// TIA Portal project "ROLLINGMILLPLC" (V16)

(* hardware
DEVICE "S71500/ET200MP station_1"  S7-1500 station
   slot 0: "Rail_0"  Rack  6ES7 590-1***0-0AA0
   slot 1: "PLC_1"  CPU 1518-4 PN/DP MFP  6ES7 518-4AX00-1AB0  V2.8
      slot 3: "CPU display_1"  6ES7591-1BA00-0AA0
      slot 32768: "PROFINET interface_1"  X1
         slot 32769: "Port_1"  X1 P1
         slot 32770: "Port_2"  X1 P2
      slot 33024: "PROFINET interface_2"  X2
         slot 33025: "Port_1"  X2 P1
      slot 33280: "PROFINET interface GBIT_3"  X3
         slot 33281: "Port_1"  X3 P1
      slot 33536: "DP interface_1"  X4
      slot 34817: "Virtual CP interface port_1"  Virtual CP interface port  Virtual CP interface port
DEVICE "S71500/ET200MP station_2"  S7-1500 station
   slot 0: "Rail_0"  Rack  6ES7 590-1***0-0AA0
   slot 1: "PLC_2"  CPU 1518-4 PN/DP MFP  6ES7 518-4AX00-1AB0  V2.8
      slot 3: "CPU display_1"  6ES7591-1BA00-0AA0
      slot 32768: "PROFINET interface_1"  X1
         slot 32769: "Port_1"  X1 P1
         slot 32770: "Port_2"  X1 P2
      slot 33024: "PROFINET interface_2"  X2
         slot 33025: "Port_1"  X2 P1
      slot 33280: "PROFINET interface GBIT_3"  X3
         slot 33281: "Port_1"  X3 P1
      slot 33536: "DP interface_1"  X4
      slot 34817: "Virtual CP interface port_1"  Virtual CP interface port  Virtual CP interface port
DEVICE "S71500/ET200MP station_3"  S7-1500 station
   slot 0: "Rail_0"  Rack  6ES7 590-1***0-0AA0
   slot 1: "PLC_3"  CPU 1518-4 PN/DP MFP  6ES7 518-4AX00-1AB0  V2.8
      slot 3: "CPU display_1"  6ES7591-1BA00-0AA0
      slot 32768: "PROFINET interface_1"  X1
         slot 32769: "Port_1"  X1 P1
         slot 32770: "Port_2"  X1 P2
      slot 33024: "PROFINET interface_2"  X2
         slot 33025: "Port_1"  X2 P1
      slot 33280: "PROFINET interface GBIT_3"  X3
         slot 33281: "Port_1"  X3 P1
      slot 33536: "DP interface_1"  X4
      slot 34817: "Virtual CP interface port_1"  Virtual CP interface port  Virtual CP interface port
DEVICE "HMI"  TP1500 Comfort
   slot 0: "HMI"  TP1500 Comfort  6AV2 124-0QC02-0AX0  16.0.0.0
   slot 1: "HMI_RT_2"  TP1500 Comfort  6AV2 124-0QC02-0AX0  16.0.0.0
   slot 5: "HMI.IE_CP_1"  PROFINET Interface  16.0.0.0
      slot 1: "PROFINET Interface_1"  PROFINET Interface
         slot 1: "Port_1"  Port
         slot 2: "Port_2"  Port
   slot 6: "HMI.IE_CP_2"  PROFINET Interface  16.0.0.0
      slot 1: "PROFINET Interface_GBit"  PROFINET Interface
         slot 1: "Port_1"  Port
   slot 7: "HMI.MPI/DP_CP_1"  MPI/DP Interface  16.0.0.0
*)

// ===== PLC "PLC_1"  CPU 1518-4 PN/DP MFP =====

TYPE "LQInternalModelSignals"
// This block is AUTO GENERATED - DO NOT MODIFY this block!
// Created by ODK_CodeGenerator version 205.100.101.18
// at Fri August 27 01:27:48 2021
// ********************************************************
   STRUCT
      Controlinput : Array[0..1] of LReal;
      Feedback : Array[0..4] of LReal;
      LQ_Refthickness : LReal;
      LQ_Refrollingforce : LReal;
   END_STRUCT;
END_TYPE

TYPE "LQParams"
// This block is AUTO GENERATED - DO NOT MODIFY this block!
// Created by ODK_CodeGenerator version 205.100.101.18
// at Mon August 30 17:02:50 2021
// ********************************************************
   STRUCT
      Lr : Array[0..3] of LReal;   // [LQ Controller 1/Gain Lr]:LQ_P.Lr
      Ly : Array[0..9] of LReal;   // [LQ Controller 1/Gain Ly]:LQ_P.Ly
   END_STRUCT;
   // Lr[0] := 0.013106;
   // Lr[1] := 0.0;
   // Lr[2] := 0.0;
   // Lr[3] := 3.112673;
   // Ly[0] := 0.0;
   // Ly[1] := 0.0;
   // Ly[2] := 0.0;
   // Ly[3] := 0.0;
   // Ly[4] := 0.011684;
   // Ly[5] := 0.0;
   // Ly[6] := 3.8E-05;
   // Ly[7] := 0.0;
   // Ly[8] := 0.0;
   // Ly[9] := 3.112673;
END_TYPE

DATA_BLOCK "LQ_GlobalData"   // DB1
{ S7_Optimized_Access := 'TRUE' }
VERSION : 0.1
   VAR
      Parameters : Struct
         thicknes : LReal;
         force : LReal;
      END_STRUCT;
      Feedback : Array[0..4] of LReal;
      Controlinput : Struct
         xv : LReal;
         fx : LReal;
      END_STRUCT;
      InternalModelSignals : "LQInternalModelSignals";
   END_VAR
   VAR RETAIN
      Param : "LQParams";
   END_VAR
BEGIN
END_DATA_BLOCK

DATA_BLOCK "gDB_SWV_Interface"   // DB2
{ S7_Optimized_Access := 'TRUE' }
VERSION : 0.1
// stored: InstanceOfName LQWebReadWrite
"LQWebReadWrite"
BEGIN
END_DATA_BLOCK

DATA_BLOCK "LQ_Unload_DB"   // DB3
{ S7_Optimized_Access := 'TRUE' }
VERSION : 0.1
// stored: InstanceOfName LQ_Unload
"LQ_Unload"
BEGIN
END_DATA_BLOCK

DATA_BLOCK "LQ_Load_DB"   // DB4
{ S7_Optimized_Access := 'TRUE' }
VERSION : 0.1
// stored: InstanceOfName LQ_Load
"LQ_Load"
BEGIN
END_DATA_BLOCK

DATA_BLOCK "LQOneStep_DB"   // DB5
{ S7_Optimized_Access := 'TRUE' }
VERSION : 0.1
// stored: InstanceOfName LQOneStep
"LQOneStep"
BEGIN
END_DATA_BLOCK

DATA_BLOCK "LQReadWriteParameters_DB"   // DB6
{ S7_Optimized_Access := 'TRUE' }
VERSION : 0.1
// stored: InstanceOfName LQReadWriteParameters
"LQReadWriteParameters"
BEGIN
END_DATA_BLOCK

DATA_BLOCK "OpcInterface"   // DB7
{ S7_Optimized_Access := 'TRUE' }
VERSION : 0.1
   VAR
      Feedback : Array[0..4] of LReal;
      Controlinput : Struct
         xv : LReal;
         fx : LReal;
      END_STRUCT;
   END_VAR
BEGIN
END_DATA_BLOCK

FUNCTION_BLOCK "LQ_Load"   // FB1, SCL
{ S7_Optimized_Access := 'TRUE' }
VERSION : 0.1
// This block is AUTO GENERATED - DO NOT MODIFY this block!
// Created by ODK_CodeGenerator version 2.5.1
// at Fri August 27 01:27:48 2021
// max. number of parallel calls into this ODK application is: 1
// *************************************************************
   VAR_INPUT
      REQ : Bool;
   END_VAR
   VAR_OUTPUT
      DONE : Bool;
      BUSY : Bool;
      ERROR : Bool;
      STATUS : Int;
   END_VAR
   VAR
      ODK_Load_Instance : ODK_Load;
      _odk_internal_LIBRARY_NAME : String := '<rt>LQ_ODK.so';
   END_VAR
   VAR CONSTANT
      _odk_internal_INSTANCE_ID : UDInt := 2_165_467_194;
   END_VAR
BEGIN
   //
   // DO NOT CHANGE BELOW OF THIS LINE !!
   // This is an automatic generated block by the
   // SIMATIC ODK 1500S V2.5.1
   // DO NOT CHANGE !!
   //
   #ODK_Load_Instance(REQ := #REQ,
                      LIBRARY_NAME := #_odk_internal_LIBRARY_NAME,
                      INSTANCE_ID := #_odk_internal_INSTANCE_ID,
                      DONE => #DONE,
                      BUSY => #BUSY,
                      ERROR => #ERROR,
                      STATUS => #STATUS);
   //
   // DO NOT CHANGE !!
   // This is an automatic generated block by the
   // SIMATIC ODK 1500S V2.5.1
   // DO NOT CHANGE ABOVE OF THIS LINE !!
   //
END_FUNCTION_BLOCK

FUNCTION_BLOCK "LQ_Unload"   // FB2, SCL
{ S7_Optimized_Access := 'TRUE' }
VERSION : 0.1
// This block is AUTO GENERATED - DO NOT MODIFY this block!
// Created by ODK_CodeGenerator version 205.100.101.18
// at Fri August 27 01:27:48 2021
// max. number of parallel calls into this ODK application is: 1
// *************************************************************
   VAR_INPUT
      REQ : Bool;
   END_VAR
   VAR_OUTPUT
      DONE : Bool;
      BUSY : Bool;
      ERROR : Bool;
      STATUS : Int;
   END_VAR
   VAR
      ODK_Unld_Instance : ODK_Unld;
   END_VAR
   VAR CONSTANT
      _odk_internal_INSTANCE_ID : UDInt := 2_165_467_194;
   END_VAR
BEGIN
   //
   // DO NOT CHANGE BELOW OF THIS LINE !!
   // This is an automatic generated block by the
   // SIMATIC ODK 1500S V2.5.1
   // DO NOT CHANGE !!
   //
   #ODK_Unld_Instance(REQ := #REQ,
                      INSTANCE_ID := #_odk_internal_INSTANCE_ID,
                      DONE => #DONE,
                      BUSY => #BUSY,
                      ERROR => #ERROR,
                      STATUS => #STATUS);
   //
   // DO NOT CHANGE !!
   // This is an automatic generated block by the
   // SIMATIC ODK 1500S V2.5.1
   // DO NOT CHANGE ABOVE OF THIS LINE !!
   //
END_FUNCTION_BLOCK

FUNCTION_BLOCK "LQOneStep"   // FB3, SCL
{ S7_Optimized_Access := 'TRUE' }
VERSION : 0.1
// This block is AUTO GENERATED - DO NOT MODIFY this block!
// Created by ODK_CodeGenerator version 205.100.101.18
// at Fri August 27 01:27:48 2021
// max. number of parallel calls into this ODK application is: 1
// *************************************************************
//  This is generated by Target 1500S for Simulink
//  Model name:                  LQ
//  Model version:               1.16
//                 
//  ODK 1500S version:           V2.5
//  Target 1500S version:        V4.0         
//  MATLAB version:              9.9 (R2020b) 29-Jul-2020
//  Simulink version:            10.2 (R2020b) 29-Jul-2020
//  MATLAB Coder version:        5.1 (R2020b) 29-Jul-2020
//  Simulink Coder version:      9.4 (R2020b) 29-Jul-2020
//  
//  ***Model details***
//  Step Size:                   0.01
//  Default parameter behaviour: Tunable
//  External Mode:               Off
//  
//  ***ODK 1500S details***  
//  Heap Size:                   32k
//  Max Block Size:              1024
//  Size of thread stack:        32k
//  SyncCallParallelCount:       1(max. number of parallel calls into this ODK application)
//  ********************************************************
   VAR_INPUT
      Feedback : Array[0..4] of LReal;
      Refthickness : LReal;
      Refrollingforce : LReal;
   END_VAR
   VAR_OUTPUT
      STATUS : Int := 0;
      xv : LReal;
      fx : LReal;
      internalSignals : "LQInternalModelSignals";
   END_VAR
   VAR
      _odk_internal_Last_REQ : Bool := FALSE;
      _odk_internal_Last_BUSY : Bool := FALSE;
      _odk_internal_IN_BUFFER : Array[0..55] of Byte;
      _odk_internal_OUT_BUFFER : Array[0..87] of Byte;
   END_VAR
   VAR_TEMP
      _odk_internal_pos : DInt;
      _odk_internal_err : Int;
      _odk_internal_i : Int;
   END_VAR
   VAR CONSTANT
      _odk_internal_INSTANCE_ID : UDInt := 2_165_467_194;
      _odk_internal_COMMAND : UDInt := 295_977_560;
   END_VAR
BEGIN
   //
   // DO NOT CHANGE BELOW OF THIS LINE !!
   // This is an automatic generated block by the
   // SIMATIC ODK 1500S V2.5.1
   // DO NOT CHANGE !!
   //
   // This is generated by Target 1500S for Simulink
   // Model name:                  LQ
   // Model version:               1.16
   //                
   // ODK 1500S version:           V2.5
   // Target 1500S version:        V4.0         
   // MATLAB version:              9.9 (R2020b) 29-Jul-2020
   // Simulink version:            10.2 (R2020b) 29-Jul-2020
   // MATLAB Coder version:        5.1 (R2020b) 29-Jul-2020
   // Simulink Coder version:      9.4 (R2020b) 29-Jul-2020
   // 
   // ***Model details***
   // Step Size:                   0.01
   // Default parameter behaviour: Tunable
   // External Mode:               Off
   // 
   // ***ODK 1500S details***  
   // Heap Size:                   32k
   // Max Block Size:              1024
   // Size of thread stack:        32k
   // SyncCallParallelCount:       1(max. number of parallel calls into this ODK application)
   // ********************************************************
   // 
   #_odk_internal_pos := 0;
   FOR #_odk_internal_i := 0 TO 4 DO
       #_odk_internal_err := WRITE_LITTLE(src_variable := #Feedback[#_odk_internal_i], dest_array := #_odk_internal_IN_BUFFER, pos := #_odk_internal_pos);
   END_FOR;
   #_odk_internal_err := WRITE_LITTLE(src_variable := #Refthickness, dest_array := #_odk_internal_IN_BUFFER, pos := #_odk_internal_pos);
   #_odk_internal_err := WRITE_LITTLE(src_variable := #Refrollingforce, dest_array := #_odk_internal_IN_BUFFER, pos := #_odk_internal_pos);
   #STATUS := ODK_ExcS(INSTANCE_ID := #_odk_internal_INSTANCE_ID,
                       COMMAND := #_odk_internal_COMMAND,
                       IN_DATA := #_odk_internal_IN_BUFFER,
                       INOUT_DATA := null,
                       OUT_DATA := #_odk_internal_OUT_BUFFER
   );
   IF INT_TO_UINT(#STATUS) < 16#7000 THEN
       #_odk_internal_pos := 0;
       #_odk_internal_err := READ_LITTLE(dest_Variable => #xv, src_array := #_odk_internal_OUT_BUFFER, pos := #_odk_internal_pos);
       #_odk_internal_err := READ_LITTLE(dest_Variable => #fx, src_array := #_odk_internal_OUT_BUFFER, pos := #_odk_internal_pos);
       FOR #_odk_internal_i := 0 TO 1 DO
           #_odk_internal_err := READ_LITTLE(dest_Variable => #internalSignals.#Controlinput[#_odk_internal_i], src_array := #_odk_internal_OUT_BUFFER, pos := #_odk_internal_pos);
       END_FOR;
       FOR #_odk_internal_i := 0 TO 4 DO
           #_odk_internal_err := READ_LITTLE(dest_Variable => #internalSignals.#Feedback[#_odk_internal_i], src_array := #_odk_internal_OUT_BUFFER, pos := #_odk_internal_pos);
       END_FOR;
       #_odk_internal_err := READ_LITTLE(dest_Variable => #internalSignals.#LQ_Refthickness, src_array := #_odk_internal_OUT_BUFFER, pos := #_odk_internal_pos);
       #_odk_internal_err := READ_LITTLE(dest_Variable => #internalSignals.#LQ_Refrollingforce, src_array := #_odk_internal_OUT_BUFFER, pos := #_odk_internal_pos);
   END_IF;
   //
   // DO NOT CHANGE !!
   // This is an automatic generated block by the
   // SIMATIC ODK 1500S V2.5.1
   // DO NOT CHANGE ABOVE OF THIS LINE !!
   //
END_FUNCTION_BLOCK

FUNCTION_BLOCK "LQReadWriteParameters"   // FB4, SCL
{ S7_Optimized_Access := 'TRUE' }
VERSION : 0.1
// This block is AUTO GENERATED - DO NOT MODIFY this block!
// Created by ODK_CodeGenerator version 205.100.101.18
// at Fri August 27 01:27:49 2021
// max. number of parallel calls into this ODK application is: 1
// *************************************************************
//  This is generated by Target 1500S for Simulink
//  Model name:                  LQ
//  Model version:               1.16
//                 
//  ODK 1500S version:           V2.5
//  Target 1500S version:        V4.0         
//  MATLAB version:              9.9 (R2020b) 29-Jul-2020
//  Simulink version:            10.2 (R2020b) 29-Jul-2020
//  MATLAB Coder version:        5.1 (R2020b) 29-Jul-2020
//  Simulink Coder version:      9.4 (R2020b) 29-Jul-2020
//  
//  ***Model details***
//  Step Size:                   0.01
//  Default parameter behaviour: Tunable
//  External Mode:               Off
//  
//  ***ODK 1500S details***  
//  Heap Size:                   32k
//  Max Block Size:              1024
//  Size of thread stack:        32k
//  SyncCallParallelCount:       1(max. number of parallel calls into this ODK application)
//  ********************************************************
//  
//  Call this function to read or write parameters from/to Simulink Model.
//  Set write[IN] parameter to TRUE in order to write and set FALSE to read parameters
   VAR_INPUT
      write : Bool;
   END_VAR
   VAR_OUTPUT
      STATUS : Int := 0;
   END_VAR
   VAR_IN_OUT
      inOutParams : "LQParams";
   END_VAR
   VAR
      _odk_internal_Last_REQ : Bool := FALSE;
      _odk_internal_Last_BUSY : Bool := FALSE;
      _odk_internal_IN_BUFFER : Array[0..0] of Byte;
      _odk_internal_INOUT_BUFFER : Array[0..111] of Byte;
   END_VAR
   VAR_TEMP
      _odk_internal_pos : DInt;
      _odk_internal_err : Int;
      _odk_internal_i : Int;
   END_VAR
   VAR CONSTANT
      _odk_internal_INSTANCE_ID : UDInt := 2_165_467_194;
      _odk_internal_COMMAND : UDInt := 2_137_970_399;
   END_VAR
BEGIN
   //
   // DO NOT CHANGE BELOW OF THIS LINE !!
   // This is an automatic generated block by the
   // SIMATIC ODK 1500S V2.5.1
   // DO NOT CHANGE !!
   //
   // This is generated by Target 1500S for Simulink
   // Model name:                  LQ
   // Model version:               1.16
   //                
   // ODK 1500S version:           V2.5
   // Target 1500S version:        V4.0         
   // MATLAB version:              9.9 (R2020b) 29-Jul-2020
   // Simulink version:            10.2 (R2020b) 29-Jul-2020
   // MATLAB Coder version:        5.1 (R2020b) 29-Jul-2020
   // Simulink Coder version:      9.4 (R2020b) 29-Jul-2020
   // 
   // ***Model details***
   // Step Size:                   0.01
   // Default parameter behaviour: Tunable
   // External Mode:               Off
   // 
   // ***ODK 1500S details***  
   // Heap Size:                   32k
   // Max Block Size:              1024
   // Size of thread stack:        32k
   // SyncCallParallelCount:       1(max. number of parallel calls into this ODK application)
   // ********************************************************
   // 
   // Call this function to read or write parameters from/to Simulink Model.
   // Set write[IN] parameter to TRUE in order to write and set FALSE to read parameters
   #_odk_internal_pos := 0;
   IF (True = #write) THEN
       #_odk_internal_IN_BUFFER[#_odk_internal_pos] := BYTE#1;
   ELSE
       #_odk_internal_IN_BUFFER[#_odk_internal_pos] := BYTE#0;
   END_IF;
   #_odk_internal_pos := #_odk_internal_pos + 1;
   #_odk_internal_pos := 0;
   FOR #_odk_internal_i := 0 TO 3 DO
       #_odk_internal_err := WRITE_LITTLE(src_variable := #inOutParams.#Lr[#_odk_internal_i], dest_array := #_odk_internal_INOUT_BUFFER, pos := #_odk_internal_pos);
   END_FOR;
   FOR #_odk_internal_i := 0 TO 9 DO
       #_odk_internal_err := WRITE_LITTLE(src_variable := #inOutParams.#Ly[#_odk_internal_i], dest_array := #_odk_internal_INOUT_BUFFER, pos := #_odk_internal_pos);
   END_FOR;
   #STATUS := ODK_ExcS(INSTANCE_ID := #_odk_internal_INSTANCE_ID,
                       COMMAND := #_odk_internal_COMMAND,
                       IN_DATA := #_odk_internal_IN_BUFFER,
                       INOUT_DATA := #_odk_internal_INOUT_BUFFER,
                       OUT_DATA := null);
   IF INT_TO_UINT(#STATUS) < 16#7000 THEN
       #_odk_internal_pos := 0;
       FOR #_odk_internal_i := 0 TO 3 DO
           #_odk_internal_err := READ_LITTLE(dest_Variable => #inOutParams.#Lr[#_odk_internal_i], src_array := #_odk_internal_INOUT_BUFFER, pos := #_odk_internal_pos);
       END_FOR;
       FOR #_odk_internal_i := 0 TO 9 DO
           #_odk_internal_err := READ_LITTLE(dest_Variable => #inOutParams.#Ly[#_odk_internal_i], src_array := #_odk_internal_INOUT_BUFFER, pos := #_odk_internal_pos);
       END_FOR;
   END_IF;
   //
   // DO NOT CHANGE !!
   // This is an automatic generated block by the
   // SIMATIC ODK 1500S V2.5.1
   // DO NOT CHANGE ABOVE OF THIS LINE !!
   //
END_FUNCTION_BLOCK

FUNCTION_BLOCK "LQWebReadWrite"   // FB5, SCL
{ S7_Optimized_Access := 'TRUE' }
VERSION : 0.1
// This block is AUTO GENERATED - DO NOT MODIFY this block!
// Created by Target 1500S version 0
// at 0 
// ********************************************************
//  This is generated by Target 1500S for Simulink
//  Model name:                  LQ
//  Model version:               1.16
//                
//  ODK 1500S version:           V2.5
//  Target 1500S version:        V4.0         
//  MATLAB version:              9.9 (R2020b) 29-Jul-2020
//  Simulink version:            10.2 (R2020b) 29-Jul-2020
//  MATLAB Coder version:        5.1 (R2020b) 29-Jul-2020
//  Simulink Coder version:      9.4 (R2020b) 29-Jul-2020
// 
//  ***Model details***
//  Step Size:                   0.01
//  Default parameter behaviour: Tunable 
//  External Mode:               Off
//  ***ODK 1500S details***  
//  Heap Size:                   32k
//  Max Block Size:              1024
//  Size of thread stack:        32k
//  SyncCallParallelCount:       1(max. number of parallel calls into this ODK application)
//  ********************************************************
// Call this FB to establish a connection to user defined Web page.
   VAR_INPUT
      InternalSignals : "LQInternalModelSignals";
      CTRL_DB : DB_WWW;
   END_VAR
   VAR_IN_OUT
      Params : "LQParams";
   END_VAR
   VAR
      TestPointedSignals : "LQInternalModelSignals";
      Parameter : "LQParams";
      RWParams_Instance : "LQReadWriteParameters";
      Write : Int := 0;
      RunTime : LReal;
   END_VAR
   VAR_TEMP
      ret : Int;
   END_VAR
BEGIN
   // This is generated by Target 1500S for Simulink
   // Model name:                  LQ
   // Model version:               1.16
   //               
   // ODK 1500S version:           V2.5
   // Target 1500S version:        V4.0         
   // MATLAB version:              9.9 (R2020b) 29-Jul-2020
   // Simulink version:            10.2 (R2020b) 29-Jul-2020
   // MATLAB Coder version:        5.1 (R2020b) 29-Jul-2020
   // Simulink Coder version:      9.4 (R2020b) 29-Jul-2020
   //
   // ***Model details***
   // Step Size:                   0.01
   // Default parameter behaviour: Tunable 
   // External Mode:               Off
   // ***ODK 1500S details***  
   // Heap Size:                   32k
   // Max Block Size:              1024
   // Size of thread stack:        32k
   // SyncCallParallelCount:       1(max. number of parallel calls into this ODK application)
   // ********************************************************
   //Call this FB to establish a connection to user defined Web page.
   #RunTime := #RunTime + 10.0;

   #TestPointedSignals := #InternalSignals;
   CASE #Write OF
       0:
           #RWParams_Instance(write := FALSE,
                              STATUS => #RWParams_Instance.STATUS,
                              inOutParams := #Parameter);
           #Params := #Parameter;
       1:
           // Wait for parameter be updated by the Web action
           ;
       2:
           #RWParams_Instance(write := TRUE,
                              STATUS => #RWParams_Instance.STATUS,
                              inOutParams := #Parameter);
           #Params := #Parameter;
           #Write := 0;
       ELSE
           // Not possible to reach
           ;
   END_CASE;

   #ret := WWW(#CTRL_DB);
END_FUNCTION_BLOCK

ORGANIZATION_BLOCK "Main"   // OB1, LAD, ProgramCycle
TITLE = "Main Program Sweep (Cycle)"
{ S7_Optimized_Access := 'TRUE' }
VERSION : 0.1
   VAR_INPUT
      Initial_Call : Bool;   // Initial call of this OB
      Remanence : Bool;   // =True, if remanent data are available
   END_VAR
BEGIN
END_ORGANIZATION_BLOCK

ORGANIZATION_BLOCK "Cyclic interrupt"   // OB30, LAD, CyclicInterrupt
{ S7_Optimized_Access := 'TRUE' }
VERSION : 0.1
   VAR_INPUT
      Initial_Call : Bool;   // Initial call of this OB
      Event_Count : Int;   // Events discarded
   END_VAR
BEGIN

REGION Network 1 (SCL)
   "LQ_GlobalData".Feedback := "OpcInterface".Feedback;
END_REGION

REGION Network 2
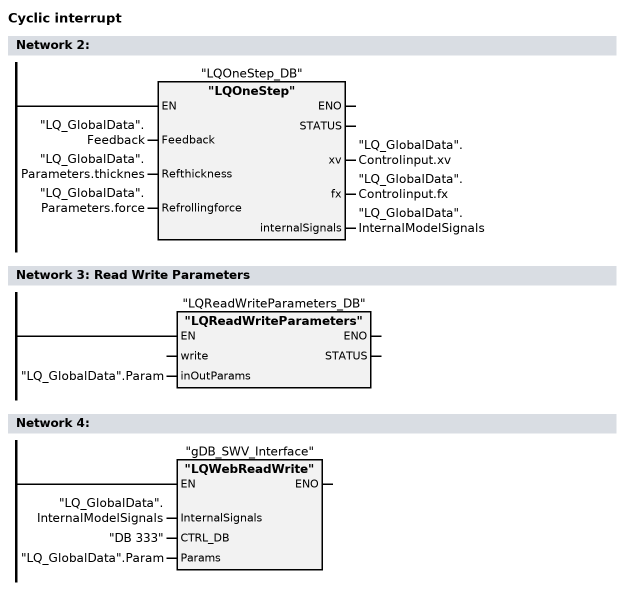
   RUNG wire#powerrail
      "LQOneStep_DB"(Feedback := "LQ_GlobalData".Feedback, Refthickness := "LQ_GlobalData".Parameters.thicknes, Refrollingforce := "LQ_GlobalData".Parameters.force, STATUS =>, xv => "LQ_GlobalData".Controlinput.xv, fx => "LQ_GlobalData".Controlinput.fx, internalSignals => "LQ_GlobalData".InternalModelSignals)
   END_RUNG
   // the same network as SCL:
   "LQOneStep_DB"(Feedback := "LQ_GlobalData".Feedback,   // "LQOneStep"
                  Refthickness := "LQ_GlobalData".Parameters.thicknes,
                  Refrollingforce := "LQ_GlobalData".Parameters.force,
                  xv => "LQ_GlobalData".Controlinput.xv,
                  fx => "LQ_GlobalData".Controlinput.fx,
                  internalSignals => "LQ_GlobalData".InternalModelSignals);
END_REGION

REGION Network 3: Read Write Parameters
   RUNG wire#powerrail
      "LQReadWriteParameters_DB"(write :=, inOutParams := "LQ_GlobalData".Param, STATUS =>)
   END_RUNG
   // the same network as SCL:
   "LQReadWriteParameters_DB"(inOutParams := "LQ_GlobalData".Param);   // "LQReadWriteParameters"
END_REGION

REGION Network 4
   RUNG wire#powerrail
      "gDB_SWV_Interface"(InternalSignals := "LQ_GlobalData".InternalModelSignals, CTRL_DB := "DB 333", Params := "LQ_GlobalData".Param)
   END_RUNG
   // the same network as SCL:
   "gDB_SWV_Interface"(InternalSignals := "LQ_GlobalData".InternalModelSignals,   // "LQWebReadWrite"
                       CTRL_DB := "DB 333",
                       Params := "LQ_GlobalData".Param);
END_REGION

REGION Network 5 (SCL)
   "OpcInterface".Controlinput.xv := "LQ_GlobalData".Controlinput.xv;
   "OpcInterface".Controlinput.fx := "LQ_GlobalData".Controlinput.fx;
END_REGION
END_ORGANIZATION_BLOCK

ORGANIZATION_BLOCK "Startup"   // OB100, LAD, Startup
TITLE = "Complete Restart"
{ S7_Optimized_Access := 'TRUE' }
VERSION : 0.1
   VAR_INPUT
      LostRetentive : Bool;   // True if retentive data are lost
      LostRTC : Bool;   // True if date and time are lost
   END_VAR
BEGIN

REGION Network 1
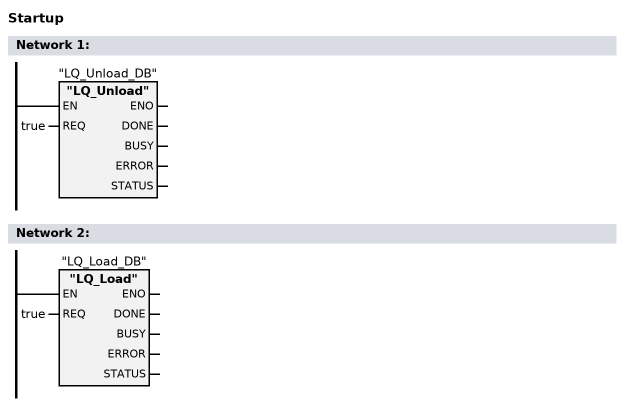
   RUNG wire#powerrail
      "LQ_Unload_DB"(REQ := true, DONE =>, BUSY =>, ERROR =>, STATUS =>)
   END_RUNG
   // the same network as SCL:
   "LQ_Unload_DB"(REQ := true);   // "LQ_Unload"
END_REGION

REGION Network 2
   RUNG wire#powerrail
      "LQ_Load_DB"(REQ := true, DONE =>, BUSY =>, ERROR =>, STATUS =>)
   END_RUNG
   // the same network as SCL:
   "LQ_Load_DB"(REQ := true);   // "LQ_Load"
END_REGION
END_ORGANIZATION_BLOCK

// ===== PLC "PLC_2"  CPU 1518-4 PN/DP MFP =====

TYPE "LQInternalModelSignals"
// This block is AUTO GENERATED - DO NOT MODIFY this block!
// Created by ODK_CodeGenerator version 205.100.101.18
// at Fri August 27 01:31:13 2021
// ********************************************************
   STRUCT
      Controlinput : Array[0..1] of LReal;
      Feedback : Array[0..4] of LReal;
      LQ_Refthickness : LReal;
      LQ_Refrollingforce : LReal;
   END_STRUCT;
END_TYPE

TYPE "LQParams"
// This block is AUTO GENERATED - DO NOT MODIFY this block!
// Created by ODK_CodeGenerator version 205.100.101.18
// at Mon August 30 17:02:50 2021
// ********************************************************
   STRUCT
      Lr : Array[0..3] of LReal;   // [LQ Controller 1/Gain Lr]:LQ_P.Lr
      Ly : Array[0..9] of LReal;   // [LQ Controller 1/Gain Ly]:LQ_P.Ly
   END_STRUCT;
   // Lr[0] := 0.013106;
   // Lr[1] := 0.0;
   // Lr[2] := 0.0;
   // Lr[3] := 3.112673;
   // Ly[0] := 0.0;
   // Ly[1] := 0.0;
   // Ly[2] := 0.0;
   // Ly[3] := 0.0;
   // Ly[4] := 0.011684;
   // Ly[5] := 0.0;
   // Ly[6] := 3.8E-05;
   // Ly[7] := 0.0;
   // Ly[8] := 0.0;
   // Ly[9] := 3.112673;
END_TYPE

DATA_BLOCK "LQ_GlobalData"   // DB1
{ S7_Optimized_Access := 'TRUE' }
VERSION : 0.1
   VAR
      Parameters : Struct
         thicknes : LReal;
         force : LReal;
      END_STRUCT;
      Feedback : Array[0..4] of LReal;
      Controlinput : Struct
         xv : LReal;
         fx : LReal;
      END_STRUCT;
      InternalModelSignals : "LQInternalModelSignals";
   END_VAR
   VAR RETAIN
      Param : "LQParams";
   END_VAR
BEGIN
END_DATA_BLOCK

DATA_BLOCK "gDB_SWV_Interface"   // DB2
{ S7_Optimized_Access := 'TRUE' }
VERSION : 0.1
// stored: InstanceOfName LQWebReadWrite
"LQWebReadWrite"
BEGIN
END_DATA_BLOCK

DATA_BLOCK "OpcInterface"   // DB3
{ S7_Optimized_Access := 'TRUE' }
VERSION : 0.1
   VAR
      Feedback : Array[0..4] of LReal;
      Controlinput : Struct
         xv : LReal;
         fx : LReal;
      END_STRUCT;
   END_VAR
BEGIN
END_DATA_BLOCK

DATA_BLOCK "LQReadWriteParameters_DB"   // DB4
{ S7_Optimized_Access := 'TRUE' }
VERSION : 0.1
// stored: InstanceOfName LQReadWriteParameters
"LQReadWriteParameters"
BEGIN
END_DATA_BLOCK

DATA_BLOCK "LQ_Unload_DB"   // DB5
{ S7_Optimized_Access := 'TRUE' }
VERSION : 0.1
// stored: InstanceOfName LQ_Unload
"LQ_Unload"
BEGIN
END_DATA_BLOCK

DATA_BLOCK "LQOneStep_DB"   // DB7
{ S7_Optimized_Access := 'TRUE' }
VERSION : 0.1
// stored: InstanceOfName LQOneStep
"LQOneStep"
BEGIN
END_DATA_BLOCK

DATA_BLOCK "LQ_Load_DB"   // DB8
{ S7_Optimized_Access := 'TRUE' }
VERSION : 0.1
// stored: InstanceOfName LQ_Load
"LQ_Load"
BEGIN
END_DATA_BLOCK

FUNCTION_BLOCK "LQ_Load"   // FB1, SCL
{ S7_Optimized_Access := 'TRUE' }
VERSION : 0.1
// This block is AUTO GENERATED - DO NOT MODIFY this block!
// Created by ODK_CodeGenerator version 2.5.1
// at Fri August 27 01:31:13 2021
// max. number of parallel calls into this ODK application is: 1
// *************************************************************
   VAR_INPUT
      REQ : Bool;
   END_VAR
   VAR_OUTPUT
      DONE : Bool;
      BUSY : Bool;
      ERROR : Bool;
      STATUS : Int;
   END_VAR
   VAR
      ODK_Load_Instance : ODK_Load;
      _odk_internal_LIBRARY_NAME : String := '<rt>LQ_ODK.so';
   END_VAR
   VAR CONSTANT
      _odk_internal_INSTANCE_ID : UDInt := 2_363_350_554;
   END_VAR
BEGIN
   //
   // DO NOT CHANGE BELOW OF THIS LINE !!
   // This is an automatic generated block by the
   // SIMATIC ODK 1500S V2.5.1
   // DO NOT CHANGE !!
   //
   #ODK_Load_Instance(REQ := #REQ,
                      LIBRARY_NAME := #_odk_internal_LIBRARY_NAME,
                      INSTANCE_ID := #_odk_internal_INSTANCE_ID,
                      DONE => #DONE,
                      BUSY => #BUSY,
                      ERROR => #ERROR,
                      STATUS => #STATUS);
   //
   // DO NOT CHANGE !!
   // This is an automatic generated block by the
   // SIMATIC ODK 1500S V2.5.1
   // DO NOT CHANGE ABOVE OF THIS LINE !!
   //
END_FUNCTION_BLOCK

FUNCTION_BLOCK "LQ_Unload"   // FB2, SCL
{ S7_Optimized_Access := 'TRUE' }
VERSION : 0.1
// This block is AUTO GENERATED - DO NOT MODIFY this block!
// Created by ODK_CodeGenerator version 205.100.101.18
// at Fri August 27 01:31:13 2021
// max. number of parallel calls into this ODK application is: 1
// *************************************************************
   VAR_INPUT
      REQ : Bool;
   END_VAR
   VAR_OUTPUT
      DONE : Bool;
      BUSY : Bool;
      ERROR : Bool;
      STATUS : Int;
   END_VAR
   VAR
      ODK_Unld_Instance : ODK_Unld;
   END_VAR
   VAR CONSTANT
      _odk_internal_INSTANCE_ID : UDInt := 2_363_350_554;
   END_VAR
BEGIN
   //
   // DO NOT CHANGE BELOW OF THIS LINE !!
   // This is an automatic generated block by the
   // SIMATIC ODK 1500S V2.5.1
   // DO NOT CHANGE !!
   //
   #ODK_Unld_Instance(REQ := #REQ,
                      INSTANCE_ID := #_odk_internal_INSTANCE_ID,
                      DONE => #DONE,
                      BUSY => #BUSY,
                      ERROR => #ERROR,
                      STATUS => #STATUS);
   //
   // DO NOT CHANGE !!
   // This is an automatic generated block by the
   // SIMATIC ODK 1500S V2.5.1
   // DO NOT CHANGE ABOVE OF THIS LINE !!
   //
END_FUNCTION_BLOCK

FUNCTION_BLOCK "LQOneStep"   // FB3, SCL
{ S7_Optimized_Access := 'TRUE' }
VERSION : 0.1
// This block is AUTO GENERATED - DO NOT MODIFY this block!
// Created by ODK_CodeGenerator version 205.100.101.18
// at Fri August 27 01:31:13 2021
// max. number of parallel calls into this ODK application is: 1
// *************************************************************
//  This is generated by Target 1500S for Simulink
//  Model name:                  LQ
//  Model version:               1.16
//                 
//  ODK 1500S version:           V2.5
//  Target 1500S version:        V4.0         
//  MATLAB version:              9.9 (R2020b) 29-Jul-2020
//  Simulink version:            10.2 (R2020b) 29-Jul-2020
//  MATLAB Coder version:        5.1 (R2020b) 29-Jul-2020
//  Simulink Coder version:      9.4 (R2020b) 29-Jul-2020
//  
//  ***Model details***
//  Step Size:                   0.01
//  Default parameter behaviour: Tunable
//  External Mode:               Off
//  
//  ***ODK 1500S details***  
//  Heap Size:                   32k
//  Max Block Size:              1024
//  Size of thread stack:        32k
//  SyncCallParallelCount:       1(max. number of parallel calls into this ODK application)
//  ********************************************************
   VAR_INPUT
      Feedback : Array[0..4] of LReal;
      Refthickness : LReal;
      Refrollingforce : LReal;
   END_VAR
   VAR_OUTPUT
      STATUS : Int := 0;
      xv : LReal;
      fx : LReal;
      internalSignals : "LQInternalModelSignals";
   END_VAR
   VAR
      _odk_internal_Last_REQ : Bool := FALSE;
      _odk_internal_Last_BUSY : Bool := FALSE;
      _odk_internal_IN_BUFFER : Array[0..55] of Byte;
      _odk_internal_OUT_BUFFER : Array[0..87] of Byte;
   END_VAR
   VAR_TEMP
      _odk_internal_pos : DInt;
      _odk_internal_err : Int;
      _odk_internal_i : Int;
   END_VAR
   VAR CONSTANT
      _odk_internal_INSTANCE_ID : UDInt := 2_363_350_554;
      _odk_internal_COMMAND : UDInt := 295_977_560;
   END_VAR
BEGIN
   //
   // DO NOT CHANGE BELOW OF THIS LINE !!
   // This is an automatic generated block by the
   // SIMATIC ODK 1500S V2.5.1
   // DO NOT CHANGE !!
   //
   // This is generated by Target 1500S for Simulink
   // Model name:                  LQ
   // Model version:               1.16
   //                
   // ODK 1500S version:           V2.5
   // Target 1500S version:        V4.0         
   // MATLAB version:              9.9 (R2020b) 29-Jul-2020
   // Simulink version:            10.2 (R2020b) 29-Jul-2020
   // MATLAB Coder version:        5.1 (R2020b) 29-Jul-2020
   // Simulink Coder version:      9.4 (R2020b) 29-Jul-2020
   // 
   // ***Model details***
   // Step Size:                   0.01
   // Default parameter behaviour: Tunable
   // External Mode:               Off
   // 
   // ***ODK 1500S details***  
   // Heap Size:                   32k
   // Max Block Size:              1024
   // Size of thread stack:        32k
   // SyncCallParallelCount:       1(max. number of parallel calls into this ODK application)
   // ********************************************************
   // 
   #_odk_internal_pos := 0;
   FOR #_odk_internal_i := 0 TO 4 DO
       #_odk_internal_err := WRITE_LITTLE(src_variable := #Feedback[#_odk_internal_i], dest_array := #_odk_internal_IN_BUFFER, pos := #_odk_internal_pos);
   END_FOR;
   #_odk_internal_err := WRITE_LITTLE(src_variable := #Refthickness, dest_array := #_odk_internal_IN_BUFFER, pos := #_odk_internal_pos);
   #_odk_internal_err := WRITE_LITTLE(src_variable := #Refrollingforce, dest_array := #_odk_internal_IN_BUFFER, pos := #_odk_internal_pos);
   #STATUS := ODK_ExcS(INSTANCE_ID := #_odk_internal_INSTANCE_ID,
                       COMMAND := #_odk_internal_COMMAND,
                       IN_DATA := #_odk_internal_IN_BUFFER,
                       INOUT_DATA := null,
                       OUT_DATA := #_odk_internal_OUT_BUFFER
   );
   IF INT_TO_UINT(#STATUS) < 16#7000 THEN
       #_odk_internal_pos := 0;
       #_odk_internal_err := READ_LITTLE(dest_Variable => #xv, src_array := #_odk_internal_OUT_BUFFER, pos := #_odk_internal_pos);
       #_odk_internal_err := READ_LITTLE(dest_Variable => #fx, src_array := #_odk_internal_OUT_BUFFER, pos := #_odk_internal_pos);
       FOR #_odk_internal_i := 0 TO 1 DO
           #_odk_internal_err := READ_LITTLE(dest_Variable => #internalSignals.#Controlinput[#_odk_internal_i], src_array := #_odk_internal_OUT_BUFFER, pos := #_odk_internal_pos);
       END_FOR;
       FOR #_odk_internal_i := 0 TO 4 DO
           #_odk_internal_err := READ_LITTLE(dest_Variable => #internalSignals.#Feedback[#_odk_internal_i], src_array := #_odk_internal_OUT_BUFFER, pos := #_odk_internal_pos);
       END_FOR;
       #_odk_internal_err := READ_LITTLE(dest_Variable => #internalSignals.#LQ_Refthickness, src_array := #_odk_internal_OUT_BUFFER, pos := #_odk_internal_pos);
       #_odk_internal_err := READ_LITTLE(dest_Variable => #internalSignals.#LQ_Refrollingforce, src_array := #_odk_internal_OUT_BUFFER, pos := #_odk_internal_pos);
   END_IF;
   //
   // DO NOT CHANGE !!
   // This is an automatic generated block by the
   // SIMATIC ODK 1500S V2.5.1
   // DO NOT CHANGE ABOVE OF THIS LINE !!
   //
END_FUNCTION_BLOCK

FUNCTION_BLOCK "LQReadWriteParameters"   // FB4, SCL
{ S7_Optimized_Access := 'TRUE' }
VERSION : 0.1
// This block is AUTO GENERATED - DO NOT MODIFY this block!
// Created by ODK_CodeGenerator version 205.100.101.18
// at Fri August 27 01:31:13 2021
// max. number of parallel calls into this ODK application is: 1
// *************************************************************
//  This is generated by Target 1500S for Simulink
//  Model name:                  LQ
//  Model version:               1.16
//                 
//  ODK 1500S version:           V2.5
//  Target 1500S version:        V4.0         
//  MATLAB version:              9.9 (R2020b) 29-Jul-2020
//  Simulink version:            10.2 (R2020b) 29-Jul-2020
//  MATLAB Coder version:        5.1 (R2020b) 29-Jul-2020
//  Simulink Coder version:      9.4 (R2020b) 29-Jul-2020
//  
//  ***Model details***
//  Step Size:                   0.01
//  Default parameter behaviour: Tunable
//  External Mode:               Off
//  
//  ***ODK 1500S details***  
//  Heap Size:                   32k
//  Max Block Size:              1024
//  Size of thread stack:        32k
//  SyncCallParallelCount:       1(max. number of parallel calls into this ODK application)
//  ********************************************************
//  
//  Call this function to read or write parameters from/to Simulink Model.
//  Set write[IN] parameter to TRUE in order to write and set FALSE to read parameters
   VAR_INPUT
      write : Bool;
   END_VAR
   VAR_OUTPUT
      STATUS : Int := 0;
   END_VAR
   VAR_IN_OUT
      inOutParams : "LQParams";
   END_VAR
   VAR
      _odk_internal_Last_REQ : Bool := FALSE;
      _odk_internal_Last_BUSY : Bool := FALSE;
      _odk_internal_IN_BUFFER : Array[0..0] of Byte;
      _odk_internal_INOUT_BUFFER : Array[0..111] of Byte;
   END_VAR
   VAR_TEMP
      _odk_internal_pos : DInt;
      _odk_internal_err : Int;
      _odk_internal_i : Int;
   END_VAR
   VAR CONSTANT
      _odk_internal_INSTANCE_ID : UDInt := 2_363_350_554;
      _odk_internal_COMMAND : UDInt := 2_137_970_399;
   END_VAR
BEGIN
   //
   // DO NOT CHANGE BELOW OF THIS LINE !!
   // This is an automatic generated block by the
   // SIMATIC ODK 1500S V2.5.1
   // DO NOT CHANGE !!
   //
   // This is generated by Target 1500S for Simulink
   // Model name:                  LQ
   // Model version:               1.16
   //                
   // ODK 1500S version:           V2.5
   // Target 1500S version:        V4.0         
   // MATLAB version:              9.9 (R2020b) 29-Jul-2020
   // Simulink version:            10.2 (R2020b) 29-Jul-2020
   // MATLAB Coder version:        5.1 (R2020b) 29-Jul-2020
   // Simulink Coder version:      9.4 (R2020b) 29-Jul-2020
   // 
   // ***Model details***
   // Step Size:                   0.01
   // Default parameter behaviour: Tunable
   // External Mode:               Off
   // 
   // ***ODK 1500S details***  
   // Heap Size:                   32k
   // Max Block Size:              1024
   // Size of thread stack:        32k
   // SyncCallParallelCount:       1(max. number of parallel calls into this ODK application)
   // ********************************************************
   // 
   // Call this function to read or write parameters from/to Simulink Model.
   // Set write[IN] parameter to TRUE in order to write and set FALSE to read parameters
   #_odk_internal_pos := 0;
   IF (True = #write) THEN
       #_odk_internal_IN_BUFFER[#_odk_internal_pos] := BYTE#1;
   ELSE
       #_odk_internal_IN_BUFFER[#_odk_internal_pos] := BYTE#0;
   END_IF;
   #_odk_internal_pos := #_odk_internal_pos + 1;
   #_odk_internal_pos := 0;
   FOR #_odk_internal_i := 0 TO 3 DO
       #_odk_internal_err := WRITE_LITTLE(src_variable := #inOutParams.#Lr[#_odk_internal_i], dest_array := #_odk_internal_INOUT_BUFFER, pos := #_odk_internal_pos);
   END_FOR;
   FOR #_odk_internal_i := 0 TO 9 DO
       #_odk_internal_err := WRITE_LITTLE(src_variable := #inOutParams.#Ly[#_odk_internal_i], dest_array := #_odk_internal_INOUT_BUFFER, pos := #_odk_internal_pos);
   END_FOR;
   #STATUS := ODK_ExcS(INSTANCE_ID := #_odk_internal_INSTANCE_ID,
                       COMMAND := #_odk_internal_COMMAND,
                       IN_DATA := #_odk_internal_IN_BUFFER,
                       INOUT_DATA := #_odk_internal_INOUT_BUFFER,
                       OUT_DATA := null);
   IF INT_TO_UINT(#STATUS) < 16#7000 THEN
       #_odk_internal_pos := 0;
       FOR #_odk_internal_i := 0 TO 3 DO
           #_odk_internal_err := READ_LITTLE(dest_Variable => #inOutParams.#Lr[#_odk_internal_i], src_array := #_odk_internal_INOUT_BUFFER, pos := #_odk_internal_pos);
       END_FOR;
       FOR #_odk_internal_i := 0 TO 9 DO
           #_odk_internal_err := READ_LITTLE(dest_Variable => #inOutParams.#Ly[#_odk_internal_i], src_array := #_odk_internal_INOUT_BUFFER, pos := #_odk_internal_pos);
       END_FOR;
   END_IF;
   //
   // DO NOT CHANGE !!
   // This is an automatic generated block by the
   // SIMATIC ODK 1500S V2.5.1
   // DO NOT CHANGE ABOVE OF THIS LINE !!
   //
END_FUNCTION_BLOCK

FUNCTION_BLOCK "LQWebReadWrite"   // FB5, SCL
{ S7_Optimized_Access := 'TRUE' }